// TIA Portal project "Vent Fan PLC" (V16) (continued)
VERSION : 0.1
   VAR_IN_OUT
      web_manual : "Station.Web_Interface.Manual.UDT";
      commands : "Drive.Commands.UDT";
   END_VAR
   VAR CONSTANT
      _RUN : String := 'run';
      _STOP : String := 'stop';
      _OVERRIDE : String := 'override';
   END_VAR
BEGIN
   "Drive.Commands.Run.Manual.Override"(web_manual := #web_manual,
                                        commands := #commands);
   IF #web_manual.mode <> #_OVERRIDE THEN
       "Drive.Commands.Run.Manual.Mode"(web_manual := #web_manual,
                                        commands := #commands);
   END_IF;
END_FUNCTION

FUNCTION "Schedule.In_Schedule" : Real   // FC11, SCL
{ S7_Optimized_Access := 'TRUE' }
VERSION : 0.1
   VAR_IN_OUT
      schedule : "Schedules.Temporal.UDT";
   END_VAR
   VAR_TEMP
      _now : DTL;
      _ret_val : Int;
      _monday : Real;
      _tuesday : Real;
      _wednesday : Real;
      _thursday : Real;
      _friday : Real;
      _saturday : Real;
      _sunday : Real;
   END_VAR
   // Ret_Val : returns speed if current time falls in any scheuled range
   VAR CONSTANT
      SUNDAY : USInt := 1;
      MONDAY : USInt := 2;
      TUESDAY : USInt := 3;
      WEDNESDAY : USInt := 4;
      THURSDAY : USInt := 5;
      FRIDAY : USInt := 6;
      SATURDAY : USInt := 7;
   END_VAR
BEGIN
   #_ret_val := RD_SYS_T(#_now);
   #_now.YEAR := 1970;
   #_now.HOUR -= 5;

   "Schedule.Encode_Weekday"(weekday := #MONDAY,
                             day_schedule := #schedule.monday);
   #_monday := "Schedule.In_Day"(day_schedule := #schedule.monday,
                                 current_time := #_now);
   IF #_monday > 0.0 THEN
       #"Schedule.In_Schedule" := #_monday;
       RETURN;
   END_IF;

   "Schedule.Encode_Weekday"(weekday := #TUESDAY,
                             day_schedule := #schedule.tuesday);
   #_tuesday := "Schedule.In_Day"(day_schedule := #schedule.tuesday,
                                  current_time := #_now);
   IF #_tuesday > 0.0 THEN
       #"Schedule.In_Schedule" := #_tuesday;
       RETURN;
   END_IF;

   "Schedule.Encode_Weekday"(weekday := #WEDNESDAY,
                             day_schedule := #schedule.wednesday);
   #_wednesday := "Schedule.In_Day"(day_schedule := #schedule.wednesday,
                                    current_time := #_now);
   IF #_wednesday > 0.0 THEN
       #"Schedule.In_Schedule" := #_wednesday;
       RETURN;
   END_IF;

   "Schedule.Encode_Weekday"(weekday := #THURSDAY,
                             day_schedule := #schedule.thursday);
   #_thursday := "Schedule.In_Day"(day_schedule := #schedule.thursday,
                                   current_time := #_now);
   IF #_thursday > 0.0 THEN
       #"Schedule.In_Schedule" := #_thursday;
       RETURN;
   END_IF;

   "Schedule.Encode_Weekday"(weekday := #FRIDAY,
                             day_schedule := #schedule.friday);
   #_friday := "Schedule.In_Day"(day_schedule := #schedule.friday,
                                 current_time := #_now);
   IF #_friday > 0.0 THEN
       #"Schedule.In_Schedule" := #_friday;
       RETURN;
   END_IF;

   "Schedule.Encode_Weekday"(weekday := #SATURDAY,
                             day_schedule := #schedule.saturday);
   #_saturday := "Schedule.In_Day"(day_schedule := #schedule.saturday,
                                   current_time := #_now);
   IF #_saturday > 0.0 THEN
       #"Schedule.In_Schedule" := #_saturday;
       RETURN;
   END_IF;

   "Schedule.Encode_Weekday"(weekday := #SUNDAY,
                             day_schedule := #schedule.sunday);
   #_sunday := "Schedule.In_Day"(day_schedule := #schedule.sunday,
                                 current_time := #_now);
   IF #_sunday > 0.0 THEN
       #"Schedule.In_Schedule" := #_sunday;
       RETURN;
   END_IF;

   #"Schedule.In_Schedule" := 0.0;
END_FUNCTION

FUNCTION "Drive.Commands.Run" : Void   // FC12, SCL
{ S7_Optimized_Access := 'TRUE' }
VERSION : 0.1
   VAR_INPUT
      current_station : Int;
      selected_station : Int;
      sensor : "Sensors.Thermal.UDT";
   END_VAR
   VAR_IN_OUT
      commands : "Drive.Commands.UDT";
      commands_manual : "Drive.Commands.UDT";
      commands_temporal : "Drive.Commands.UDT";
      commands_thermal : "Drive.Commands.UDT";
      web_manual : "Station.Web_Interface.Manual.UDT";
      thermal : "Schedules.Thermal.UDT";
      temporal : "Schedules.Temporal.UDT";
   END_VAR
BEGIN
   REGION "TEMPORAL"
       "Drive.Commands.Run.Temporal"(schedule:=#temporal,
                                     commands:=#commands_temporal);
       "Drive.Commands.Run.Temporal"(commands:=#commands_temporal,
                                     schedule:=#temporal);

   END_REGION

   REGION "THERMAL"
       "Drive.Commands.Run.Thermal"(sensor := #sensor,
                                    schedule := #thermal,
                                    commands := #commands_thermal);
   END_REGION

   REGION "MANUAL"
       IF #selected_station = #current_station THEN
           "Drive.Commands.Run.Manual"(web_manual := #web_manual,
                                       commands := #commands_manual);
       END_IF;
   END_REGION

   REGION "RESOLVE COMMANDS"
       "Drive.Commands.Run.Actual"(manual := #commands_manual,
                                   temporal := #commands_temporal,
                                   thermal := #commands_thermal,
                                   actual := #commands);
   END_REGION ;
END_FUNCTION

FUNCTION "Drive.Commands" : Void   // FC13, SCL
{ S7_Optimized_Access := 'TRUE' }
VERSION : 0.1
   VAR_INPUT
      current_station : Int;
      selected_station : Int;
      thermal_sensor : "Sensors.Thermal.UDT";
   END_VAR
   VAR_IN_OUT
      commands : "Drive.Commands.UDT";
      commands_manual : "Drive.Commands.UDT";
      commands_temporal : "Drive.Commands.UDT";
      commands_thermal : "Drive.Commands.UDT";
      manual : "Station.Web_Interface.Manual.UDT";
      thermal : "Schedules.Thermal.UDT";
      temporal : "Schedules.Temporal.UDT";
   END_VAR
BEGIN
   "Drive.Commands.Run"(current_station := #current_station,
                        selected_station := #selected_station,
                        sensor := #thermal_sensor,
                        commands := #commands,
                        commands_manual := #commands_manual,
                        commands_thermal := #commands_thermal,
                        commands_temporal := #commands_temporal,
                        web_manual := #manual,
                        thermal := #thermal,
                        temporal := #temporal);
END_FUNCTION

FUNCTION "Drive.Commands.Run.Actual" : Void   // FC14, SCL
{ S7_Optimized_Access := 'TRUE' }
VERSION : 0.1
   VAR_INPUT
      manual : "Drive.Commands.UDT";
      temporal : "Drive.Commands.UDT";
      thermal : "Drive.Commands.UDT";
   END_VAR
   VAR_IN_OUT
      actual : "Drive.Commands.UDT";
   END_VAR
BEGIN
   IF #manual.stop THEN
       #actual := #manual;
       RETURN;
   END_IF;

   IF #manual.override THEN
       #actual := #manual;
       RETURN;
   END_IF;

   IF #thermal.run THEN
       #actual := #thermal;
       RETURN;
   END_IF;

   IF #temporal.run THEN
       #actual := #temporal;
       RETURN;
   END_IF;

   #actual.speed := "Drive.Protection.Bound_Percentage"(#actual.speed);

   "Drive.Command_Stop"(#actual);
END_FUNCTION

FUNCTION "Real.Scale" : Real   // FC15, SCL
{ S7_Optimized_Access := 'TRUE' }
VERSION : 0.1
   VAR_INPUT
      x_min : Real;
      x_max : Real;
      x_actual : Real;
      y_min : Real;
      y_max : Real;
   END_VAR
BEGIN
   #"Real.Scale" := (#y_max - #y_min) / (#x_max - #x_min) * (#x_actual - #x_min) + (#y_min);
END_FUNCTION

FUNCTION "String.Split" : Void   // FC16, SCL
{ S7_Optimized_Access := 'TRUE' }
VERSION : 0.1
   VAR_INPUT
      string_in : String;
      delimeter : String;
      pointer : Int;   // pointer for recursion
   END_VAR
   VAR_IN_OUT
      sub_strings : Array[*] of String;
   END_VAR
   VAR_TEMP
      _split : String;
      _position : Int;
      _return : String;
   END_VAR
BEGIN
   REGION "GET POSITION OF DELIMETER IN STRING"
       #_position := FIND(IN1 := #string_in,
                          IN2 := #delimeter);
   END_REGION

   REGION "BASE CASE"
       IF #_position = 0 THEN
           #sub_strings[#pointer] := #string_in;
           RETURN;
       END_IF;
   END_REGION


   REGION "RECURSIVE CASE"
       #sub_strings[#pointer] := LEFT(IN := #string_in, L := #_position - 1);
       "String.Split"(string_in := RIGHT(IN := #string_in, L := LEN(#string_in) - #_position),
                      delimeter := #delimeter,
                      "pointer" := #pointer + 1,
                      sub_strings := #sub_strings);
   END_REGION
END_FUNCTION

FUNCTION "Schedule.Temporal.Clean_Data" : Void   // FC17, SCL
{ S7_Optimized_Access := 'TRUE' }
VERSION : 0.1
   VAR_IN_OUT
      schedule : "Schedules.Temporal.UDT";
   END_VAR
BEGIN
END_FUNCTION

FUNCTION "Web_Meta.Update_Temporal" : Void   // FC18, SCL
{ S7_Optimized_Access := 'TRUE' }
VERSION : 0.1
   VAR_IN_OUT
      web_schedules : "Web_Meta.Web_Interface.Schedules.Temporal.UDT";
      plc_schedules : "Schedules.Temporal.UDT";
   END_VAR
BEGIN
   IF NOT #web_schedules.new_data THEN
       RETURN;
   END_IF;

   "Web_Meta.Update_Temporal.Web_to_PLC"(web := #web_schedules,
                                         plc := #plc_schedules);
   #web_schedules.new_data := FALSE;
END_FUNCTION

FUNCTION "Web_Meta.Update_Temporal.Web_to_PLC" : Void   // FC19, SCL
{ S7_Optimized_Access := 'TRUE' }
VERSION : 0.1
   VAR_INPUT
      web : "Web_Meta.Web_Interface.Schedules.Temporal.UDT";
   END_VAR
   VAR_IN_OUT
      plc : "Schedules.Temporal.UDT";
   END_VAR
BEGIN
   "Web_Meta.Update_Temporal.Web_to_PLC.Day"(web := #web.monday,
                                             plc := #plc.monday);
   "Web_Meta.Update_Temporal.Web_to_PLC.Day"(web := #web.tuesday,
                                             plc := #plc.tuesday);
   "Web_Meta.Update_Temporal.Web_to_PLC.Day"(web := #web.wednesday,
                                             plc := #plc.wednesday);
   "Web_Meta.Update_Temporal.Web_to_PLC.Day"(web := #web.thursday,
                                             plc := #plc.thursday);
   "Web_Meta.Update_Temporal.Web_to_PLC.Day"(web := #web.friday,
                                             plc := #plc.friday);
   "Web_Meta.Update_Temporal.Web_to_PLC.Day"(web := #web.saturday,
                                             plc := #plc.saturday);
   "Web_Meta.Update_Temporal.Web_to_PLC.Day"(web := #web.sunday,
                                             plc := #plc.sunday);
END_FUNCTION

FUNCTION "Web_Meta.Update_Temporal.PLC_to_Web" : Void   // FC20, SCL
{ S7_Optimized_Access := 'TRUE' }
VERSION : 0.1
   VAR_INPUT
      plc : "Schedules.Temporal.UDT";
   END_VAR
   VAR_IN_OUT
      web : "Web_Meta.Web_Interface.Schedules.Temporal.UDT";
   END_VAR
BEGIN
   "Web_Meta.Update_Temporal.PLC_to_Web.Day"(plc := #plc.monday,
                                             web := #web.monday);
   "Web_Meta.Update_Temporal.PLC_to_Web.Day"(plc := #plc.tuesday,
                                             web := #web.tuesday);
   "Web_Meta.Update_Temporal.PLC_to_Web.Day"(plc := #plc.wednesday,
                                             web := #web.wednesday);
   "Web_Meta.Update_Temporal.PLC_to_Web.Day"(plc := #plc.thursday,
                                             web := #web.thursday);
   "Web_Meta.Update_Temporal.PLC_to_Web.Day"(plc := #plc.friday,
                                             web := #web.friday);
   "Web_Meta.Update_Temporal.PLC_to_Web.Day"(plc := #plc.saturday,
                                             web := #web.saturday);
   "Web_Meta.Update_Temporal.PLC_to_Web.Day"(plc := #plc.sunday,
                                             web := #web.sunday);
END_FUNCTION

FUNCTION "Web_Meta.Update_Temporal.PLC_to_Web.Day" : Void   // FC21, SCL
{ S7_Optimized_Access := 'TRUE' }
VERSION : 0.1
   VAR_INPUT
      plc : Array[0.."SCHEDULES_PER_DAY"] of "Schedules.Temporal.Element.UDT";
   END_VAR
   VAR_IN_OUT
      web : Array[0.."SCHEDULES_PER_DAY"] of "Web_Meta.Web_Interface.Schedules.Temporal.Element.UDT";
   END_VAR
   VAR_TEMP
      _i : Int;
   END_VAR
BEGIN
   FOR #_i := 0 TO "SCHEDULES_PER_DAY" DO
       #web[#_i].start := "Web_Meta.Update_Temporal.PLC_to_Web.Day.Element"(#plc[#_i].start);
       #web[#_i].stop := "Web_Meta.Update_Temporal.PLC_to_Web.Day.Element"(#plc[#_i].stop);
       #web[#_i].speed := #plc[#_i].speed;
   END_FOR;
END_FUNCTION

FUNCTION "Web_Meta.Update_Temporal.PLC_to_Web.Day.Element" : String   // FC22, SCL
{ S7_Optimized_Access := 'TRUE' }
VERSION : 0.1
   VAR_INPUT
      plc : "Schedules.Temporal.Element.Date_Time.UDT";
   END_VAR
   VAR_TEMP
      _ret : String;
   END_VAR
   VAR CONSTANT
      YEAR : String := '2022';
      "-" : String := '-';
   END_VAR
BEGIN
   // format --> value="2017-06-01T08:30"
   #_ret := CONCAT_STRING(IN1 := #YEAR,
                          IN2 := '-',
                          IN3 := "USInt.Convert.String.Date_with_Leading_Zeros"(#plc.month),
                          IN4 := '-',
                          IN5 := "USInt.Convert.String.Date_with_Leading_Zeros"(#plc.day),
                          IN6 := 'T',
                          IN7 := "USInt.Convert.String.Date_with_Leading_Zeros"(#plc.hour),
                          IN8 := ':',
                          IN9 := "USInt.Convert.String.Date_with_Leading_Zeros"(#plc.minute));
   #"Web_Meta.Update_Temporal.PLC_to_Web.Day.Element" := #_ret;
END_FUNCTION

FUNCTION "String.Strip Sign" : String   // FC23, SCL
{ S7_Optimized_Access := 'TRUE' }
VERSION : 0.1
   VAR_INPUT
      "string" : String;
   END_VAR
   VAR_TEMP
      Length : Int;
      "String Box" : String;
      "Test Character" : String;
   END_VAR
   VAR CONSTANT
      "+" : Char := '+';
      "-" : Char := '-';
   END_VAR
BEGIN
   #"String Box" := #string;
   #"Test Character" := LEFT_STRING(IN := #"String Box",
                                    L := 1);
   IF #"Test Character" = #"+" OR #"Test Character" = #"-" THEN
       #Length := LEN(#"String Box");
       #"String Box" := RIGHT_STRING(IN := #"String Box", L := #Length - 1);

   END_IF;
   #"String.Strip Sign" := #"String Box";
END_FUNCTION

FUNCTION "String.Trim" : String   // FC24, SCL
{ S7_Optimized_Access := 'TRUE' }
AUTHOR : Machado
FAMILY : String
VERSION : 1.0
// removes leading and trailing whitespace from input string
   VAR_INPUT
      "string" : String;
   END_VAR
   VAR_TEMP
      ret : String;
   END_VAR
   VAR CONSTANT
      space : String := ' ';
   END_VAR
BEGIN
   #ret := #string;
   WHILE LEFT(IN := #ret, L := 1) = #space DO
       #ret := RIGHT(IN := #ret, L := LEN(#ret) - 1);
   END_WHILE;
   WHILE RIGHT(IN := #ret, L := 1) = #space DO
       #ret := LEFT(IN := #ret, L := LEN(#ret) - 1);
   END_WHILE;
   #"String.Trim" := #ret;
END_FUNCTION

FUNCTION "USInt.Convert.Clean_String" : String   // FC25, SCL
{ S7_Optimized_Access := 'TRUE' }
VERSION : 0.1
   VAR_INPUT
      in : USInt;
   END_VAR
BEGIN
   #"USInt.Convert.Clean_String" := "String.Trim"("String.Strip Sign"(USINT_TO_STRING(#in)));
END_FUNCTION

FUNCTION "String.Add Leading" : String   // FC26, SCL
{ S7_Optimized_Access := 'TRUE' }
VERSION : 0.1
   VAR_INPUT
      "Leading Character" : Char;
      "Desired Length" : USInt;
      "String" : String;
   END_VAR
   VAR_TEMP
      Length : Int;
      "String Box" : String;
   END_VAR
BEGIN
   #"String Box" := #String;
   #Length := LEN(#"String Box");

   WHILE #Length < #"Desired Length" DO
       #"String Box" := CONCAT_STRING(IN1 := #"Leading Character",
                                      IN2 := #"String Box");
       #Length := LEN(#"String Box");
   END_WHILE;

   #"String.Add Leading" := #"String Box";
END_FUNCTION

FUNCTION "USInt.Convert.String.Date_with_Leading_Zeros" : String   // FC27, SCL
{ S7_Optimized_Access := 'TRUE' }
VERSION : 0.1
   VAR_INPUT
      in : USInt;
   END_VAR
BEGIN
   #"USInt.Convert.String.Date_with_Leading_Zeros" := "String.Add Leading"("Leading Character" := '0',
                                                                           "Desired Length" := 2,
                                                                           "String" := "USInt.Convert.Clean_String"(#in));
END_FUNCTION

FUNCTION "Web_Meta.Update_Temporal.Web_to_PLC.Day.Element" : "Schedules.Temporal.Element.Date_Time.UDT"   // FC28, SCL
{ S7_Optimized_Access := 'TRUE' }
VERSION : 0.1
   VAR_INPUT
      in : String;
   END_VAR
   VAR_TEMP
      _ret : "Schedules.Temporal.Element.Date_Time.UDT";
      _split_date_time : Array[0..1] of String;
      _split_date : Array[0..2] of String;
      _split_time : Array[0..1] of String;
   END_VAR
BEGIN
   // format --> value="2017-06-01T08:30"
   REGION "SPLIT INTO DATE AND TIME"
       "String.Split"(string_in := #in,
                      delimeter := 'T',
                      "pointer" := 0,
                      sub_strings := #_split_date_time);
   END_REGION

   REGION "SPLIT DATE INTO YEARS, MONTHS, AND DAYS"
       "String.Split"(string_in := #_split_date_time[0],
                      delimeter := '-',
                      "pointer" := 0,
                      sub_strings := #_split_date);
   END_REGION

   REGION "SPLIT TIME INTO HOURS AND MINUTES"
       "String.Split"(string_in := #_split_date_time[1],
                      delimeter := ':',
                      "pointer" := 0,
                      sub_strings := #_split_time);
   END_REGION

   REGION "MAP TO UDT"
       #_ret.month := STRING_TO_USINT(#_split_date[1]);
       #_ret.day := STRING_TO_USINT(#_split_date[2]);
       #_ret.hour := STRING_TO_USINT(#_split_time[0]);
       #_ret.minute := STRING_TO_USINT(#_split_time[1]);
   END_REGION

   REGION "RETURN DATA"
       #"Web_Meta.Update_Temporal.Web_to_PLC.Day.Element" := #_ret;
   END_REGION
END_FUNCTION

FUNCTION "Web_Meta.Update_Temporal.Web_to_PLC.Day" : Void   // FC29, SCL
{ S7_Optimized_Access := 'TRUE' }
VERSION : 0.1
   VAR_INPUT
      web : Array[0.."SCHEDULES_PER_DAY"] of "Web_Meta.Web_Interface.Schedules.Temporal.Element.UDT";
   END_VAR
   VAR_IN_OUT
      plc : Array[0.."SCHEDULES_PER_DAY"] of "Schedules.Temporal.Element.UDT";
   END_VAR
   VAR_TEMP
      _i : Int;
   END_VAR
BEGIN
   FOR #_i := 0 TO "SCHEDULES_PER_DAY" DO
       #plc[#_i].start := "Web_Meta.Update_Temporal.Web_to_PLC.Day.Element"(#web[#_i].start);
       #plc[#_i].stop := "Web_Meta.Update_Temporal.Web_to_PLC.Day.Element"(#web[#_i].stop);
       #plc[#_i].speed := #web[#_i].speed;
   END_FOR;
END_FUNCTION

FUNCTION "Schedule.In_Day" : Real   // FC30, SCL
{ S7_Optimized_Access := 'TRUE' }
VERSION : 0.1
   VAR_INPUT
      day_schedule : Array[0.."SCHEDULES_PER_DAY"] of "Schedules.Temporal.Element.UDT";
      current_time : DTL;
   END_VAR
   VAR_TEMP
      _i : Int;
      _speed : Real;
   END_VAR
BEGIN
   IF #current_time.WEEKDAY <> #day_schedule[0].start.weekday THEN
       #"Schedule.In_Day" := 0.0;
       RETURN;
   END_IF;
   FOR #_i := 0 TO "SCHEDULES_PER_DAY" DO
       #_speed := "Schedule.In_Window"(day := #day_schedule[#_i],
                                       now := #current_time);
       IF #_speed > 0.0 THEN
           #"Schedule.In_Day" := #_speed;
           RETURN;
       END_IF;
   END_FOR;
   #"Schedule.In_Day" := 0.0;
END_FUNCTION

FUNCTION "Schedule.In_Window" : Real   // FC31, SCL
{ S7_Optimized_Access := 'TRUE' }
VERSION : 0.1
   VAR_INPUT
      day : "Schedules.Temporal.Element.UDT";
      now : DTL;
   END_VAR
   VAR_TEMP
      _start : DTL;
      _stop : DTL;
   END_VAR
BEGIN
   #_start := "Schedule.Map.Date_Time_to_DTL"(#day.start);
   #_stop := "Schedule.Map.Date_Time_to_DTL"(#day.stop);
   IF #_start < #now AND #now < #_stop THEN
       #"Schedule.In_Window" := #day.speed;
       RETURN;
   END_IF;
   #"Schedule.In_Window" := 0.0;
END_FUNCTION

FUNCTION "Schedule.Map.Date_Time_to_DTL" : DTL   // FC32, SCL
{ S7_Optimized_Access := 'TRUE' }
VERSION : 0.1
   VAR_INPUT
      boundary : "Schedules.Temporal.Element.Date_Time.UDT";
   END_VAR
   VAR_TEMP
      _ret : DTL;
   END_VAR
BEGIN
   #_ret.MONTH := #boundary.month;
   #_ret.DAY := #boundary.day;
   #_ret.HOUR := #boundary.hour;
   #_ret.MINUTE := #boundary.minute;
   #"Schedule.Map.Date_Time_to_DTL" := #_ret;
END_FUNCTION

FUNCTION "Drive.Commands.Run.Temporal" : Void   // FC33, SCL
{ S7_Optimized_Access := 'TRUE' }
VERSION : 0.1
   VAR_IN_OUT
      commands : "Drive.Commands.UDT";
      schedule : "Schedules.Temporal.UDT";
   END_VAR
   VAR_TEMP
      _speed : Real;
   END_VAR
BEGIN
   #_speed := "Schedule.In_Schedule"(schedule:=#schedule);

   IF #_speed = 0.0 THEN
       "Drive.Command_Stop"(#commands);
       RETURN;
   END_IF;

   "Drive.Command_Run"(speed := #_speed,
                       commands := #commands);
END_FUNCTION

FUNCTION "Drive.Command_Run" : Void   // FC34, SCL
{ S7_Optimized_Access := 'TRUE' }
VERSION : 0.1
   VAR_INPUT
      speed : Real;
   END_VAR
   VAR_IN_OUT
      commands : "Drive.Commands.UDT";
   END_VAR
BEGIN
   #commands.run := TRUE;
   #commands.stop := FALSE;
   #commands.speed := #speed;
END_FUNCTION

FUNCTION "Drive.Command_Stop" : Void   // FC35, SCL
{ S7_Optimized_Access := 'TRUE' }
VERSION : 0.1
   VAR_IN_OUT
      commands : "Drive.Commands.UDT";
   END_VAR
BEGIN
   #commands.run := FALSE;
   #commands.stop := TRUE;
   #commands.speed := 0.0;
END_FUNCTION

FUNCTION "Nibble.ToString" : String   // FC36, SCL
{ S7_Optimized_Access := 'TRUE' }
VERSION : 0.1
   VAR_INPUT
      value : Byte;
   END_VAR
   VAR_TEMP
      _nibble_as_int : Int;
      _ret : String;
   END_VAR
BEGIN
   #_nibble_as_int := BYTE_TO_INT(#value);
   CASE #_nibble_as_int OF
       0..9:
           #_ret := "String.Trim"("String.Strip Sign"(INT_TO_STRING(#_nibble_as_int)));
       10:
           #_ret := 'A';
       11:
           #_ret := 'B';
       12:
           #_ret := 'C';
       13:
           #_ret := 'D';
       14:
           #_ret := 'E';
       15:
           #_ret := 'F';
   END_CASE;
   #"Nibble.ToString" := #_ret;
END_FUNCTION

FUNCTION "Byte.ToString" : String   // FC37, SCL
{ S7_Optimized_Access := 'TRUE' }
VERSION : 0.1
   VAR_INPUT
      value : Byte;
   END_VAR
   VAR_TEMP
      _low_nibble : Byte;
      _high_nibble : Byte;
   END_VAR
   VAR CONSTANT
      LOW_NIBBLE_MASK : Byte := 16#0F;
      HIGH_NIBBLE_MASK : Byte := 16#F0;
   END_VAR
BEGIN
   #_low_nibble := #value AND #LOW_NIBBLE_MASK;
   #_high_nibble := SHR_BYTE(IN := #value AND #HIGH_NIBBLE_MASK,
                             N := 4);
   #"Byte.ToString" := CONCAT_STRING(IN1 := "Nibble.ToString"(#_high_nibble),
                                     IN2 := "Nibble.ToString"(#_low_nibble));
END_FUNCTION

FUNCTION "Drive.Feedback.Speed.Percent_to_RPM" : Real   // FC38, SCL
{ S7_Optimized_Access := 'TRUE' }
VERSION : 0.1
   VAR_INPUT
      as_percent : Real;
      max_speed : Real;
   END_VAR
BEGIN
   #"Drive.Feedback.Speed.Percent_to_RPM" := "Drive.Protection.Bound_Percentage"(#as_percent/100) * #max_speed;
END_FUNCTION

FUNCTION "Drive.Protection.Bound_Percentage" : Real   // FC39, SCL
{ S7_Optimized_Access := 'TRUE' }
VERSION : 0.1
   VAR_INPUT
      value : Real;
   END_VAR
BEGIN
   IF #value > 1.0 THEN
       #"Drive.Protection.Bound_Percentage" := 1.0;
       RETURN;
   END_IF;

   IF #value < 0.0 THEN
       #"Drive.Protection.Bound_Percentage" := 0.0;
       RETURN;
   END_IF;

   #"Drive.Protection.Bound_Percentage" := #value;
END_FUNCTION

FUNCTION "Schedule.Encode_Weekday" : Void   // FC40, SCL
{ S7_Optimized_Access := 'TRUE' }
VERSION : 0.1
   VAR_INPUT
      weekday : USInt;
   END_VAR
   VAR_IN_OUT
      day_schedule : Array[0.."SCHEDULES_PER_DAY"] of "Schedules.Temporal.Element.UDT";
   END_VAR
   VAR_TEMP
      i : Int;
   END_VAR
BEGIN
   FOR #i := 0 TO "SCHEDULES_PER_DAY" DO
       #day_schedule[#i].start.weekday := #weekday;
       #day_schedule[#i].stop.weekday := #weekday;
   END_FOR;
END_FUNCTION

FUNCTION "Drive.Feedback.Speed.RPM_to_Percent" : Real   // FC41, SCL
{ S7_Optimized_Access := 'TRUE' }
VERSION : 0.1
   VAR_INPUT
      as_rpm : Real;
      max_speed : Real;
   END_VAR
BEGIN
   #"Drive.Feedback.Speed.RPM_to_Percent" := #as_rpm / #max_speed * 100.0;
END_FUNCTION

FUNCTION "Drive.Commands.Run.Manual.Override" : Void   // FC42, SCL
{ S7_Optimized_Access := 'TRUE' }
VERSION : 0.1
   VAR_IN_OUT
      web_manual : "Station.Web_Interface.Manual.UDT";
      commands : "Drive.Commands.UDT";
   END_VAR
   VAR CONSTANT
      _RUN : String := 'run';
      _STOP : String := 'stop';
      _OVERRIDE : String := 'override';
   END_VAR
BEGIN
   IF #web_manual.toggle AND #web_manual.mode = #_OVERRIDE THEN
       #web_manual.mode := #_STOP;
       #web_manual.toggle := FALSE;
       #web_manual.override := FALSE;
       #commands.override := FALSE;
       #commands.run := FALSE;
       #commands.stop := TRUE;
       #commands.speed := 0.0;
       RETURN;
   END_IF;
   IF #web_manual.override THEN
       #web_manual.mode := #_OVERRIDE;
       #commands.override := TRUE;
       #commands.run := TRUE;
       #commands.stop := FALSE;
       #commands.speed := #web_manual.command_speed;
       RETURN;
   END_IF;
   IF NOT #web_manual.override AND #web_manual.mode = #_OVERRIDE THEN
       #web_manual.mode := #_STOP;
       #commands.override := FALSE;
       #commands.run := FALSE;
       #commands.stop := TRUE;
       #commands.speed := 0.0;
   END_IF;
END_FUNCTION

FUNCTION "Drive.Commands.Run.Manual.Mode" : Void   // FC43, SCL
{ S7_Optimized_Access := 'TRUE' }
VERSION : 0.1
   VAR_IN_OUT
      web_manual : "Station.Web_Interface.Manual.UDT";
      commands : "Drive.Commands.UDT";
   END_VAR
   VAR CONSTANT
      _RUN : String := 'run';
      _STOP : String := 'stop';
   END_VAR
BEGIN
   IF NOT #web_manual.toggle THEN
       RETURN;
   END_IF;
   IF #web_manual.mode = #_RUN THEN
       #web_manual.mode := #_STOP;
       #commands.run := FALSE;
       #commands.stop := TRUE;
       #commands.speed := 0.0;
       #web_manual.toggle := FALSE;
       RETURN;
   END_IF;
   IF #web_manual.mode = #_STOP THEN
       #web_manual.mode := #_RUN;
       #commands.run := TRUE;
       #commands.stop := FALSE;
       #web_manual.toggle := FALSE;
   END_IF;
END_FUNCTION

FUNCTION "Web_Meta.Update_Manual.PLC_to_Web" : Void   // FC44, SCL
{ S7_Optimized_Access := 'TRUE' }
VERSION : 0.1
   VAR_INPUT
      station : "Station.UDT";
   END_VAR
   VAR_IN_OUT
      manual : "Station.Web_Interface.Manual.UDT";
   END_VAR
BEGIN
   #manual.command_speed := #station.drive.commands_manual.speed;
   #manual.override := #station.drive.commands_manual.override;
   IF #station.drive.commands.override THEN
       #manual.mode := 'override';
   END_IF;
   IF #station.drive.commands.run THEN
       #manual.mode := 'run';
   END_IF;
   IF #station.drive.commands.stop THEN
       #manual.mode := 'stop';
   END_IF;
END_FUNCTION

FUNCTION "Faults" : Void   // FC45, SCL
{ S7_Optimized_Access := 'TRUE' }
VERSION : 0.1
   VAR_INPUT
      fault_code : Word;
   END_VAR
   VAR_IN_OUT
      station : "Station.UDT";
   END_VAR
   VAR_TEMP
      _drive_speed : Real;
      _command_speed : Real;
      _current : Real;
   END_VAR
   VAR CONSTANT
      NO_FAULT : Word := 16#7002;
      COMM_FAULT : Word := 16#80B1;
      RED : String := 'red';
      BLUE : String := 'blue';
      YELLOW : String := 'yellow';
      GREEN : String := 'green';
   END_VAR
BEGIN
   #station.faults.fault := 'no faults';
   #station.faults.color := '';

   #_drive_speed := #station.drive.feedback.speed.me.processed;
   #_command_speed := #station.drive.commands.speed;
   #_current := #station.drive.feedback.current.me.processed;

   IF #fault_code >= #NO_FAULT THEN
       IF #fault_code <> #COMM_FAULT THEN
           #station.faults.fault := "Word.ToString"(#fault_code);
           #station.faults.color := #RED;
           RETURN;
       END_IF;
   END_IF;

   IF #_drive_speed = 0.0 THEN
       IF #_command_speed <> 0.0 THEN
           #station.faults.fault := 'stopped while commanded speed above 0.0';
           #station.faults.color := #YELLOW;
           RETURN;
       END_IF;
   END_IF;

   IF #_command_speed > 10.0 THEN
       IF #_current < 2.0 THEN
           #station.faults.fault := 'low current draw';
           #station.faults.color := #RED;
           RETURN;
       END_IF;
   END_IF;

   IF #_command_speed > 10.0 THEN
       IF #_current > 6.0 THEN
           #station.faults.fault := 'high current draw';
           #station.faults.color := #RED;
           RETURN;
       END_IF;
   END_IF;

   IF #_current > 7.0 THEN
       #station.drive.commands.speed := 0.0;
       #station.faults.fault := 'over current';
       #station.faults.color := #RED;
       RETURN;
   END_IF;

   IF #_drive_speed = 0.0 THEN
       IF #_command_speed = 0.0 THEN
           #station.faults.fault := 'drive commanded stop';
           #station.faults.color := #BLUE;
           RETURN;
       END_IF;
   END_IF;

   IF #_drive_speed > 0.9 * #_command_speed THEN
       IF #_drive_speed < 1.1 * #_command_speed THEN
           #station.faults.fault := 'no faults';
           #station.faults.color := #GREEN;
           RETURN;
       END_IF;
   END_IF;
END_FUNCTION

ORGANIZATION_BLOCK "Main"   // OB1, LAD, ProgramCycle
TITLE = "Main Program Sweep (Cycle)"
{ S7_Optimized_Access := 'TRUE' }
VERSION : 0.1
   VAR_INPUT
      Initial_Call : Bool;   // Initial call of this OB
      Remanence : Bool;   // =True, if remanent data are available
   END_VAR
   VAR_TEMP
      RET_VAL : Int;
   END_VAR
   VAR CONSTANT
      SENSOR_MAX : Word := 16#3F_FF;
      SENSOR_MIN : Word;
      THERMAL_MAX : Real := 150.0;
      THERMAL_MIN : Real;
   END_VAR
BEGIN

REGION Network 1
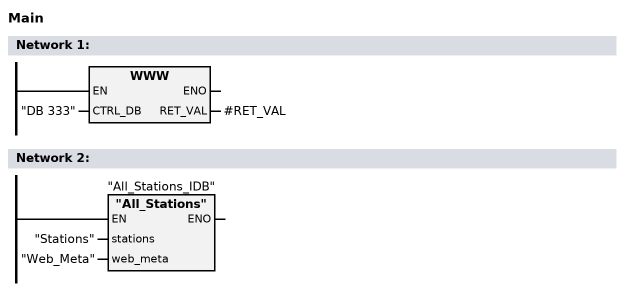
   #RET_VAL := WWW(CTRL_DB := "DB 333");
END_REGION

REGION Network 2
   RUNG wire#powerrail
      "All_Stations_IDB"(stations := "Stations", web_meta := "Web_Meta")
   END_RUNG
   // the same network as SCL:
   "All_Stations_IDB"(stations := "Stations", web_meta := "Web_Meta");   // "All_Stations"
END_REGION
END_ORGANIZATION_BLOCK

ORGANIZATION_BLOCK "Time error interrupt"   // OB80, LAD, TimeErrorInterrupt
{ S7_Optimized_Access := 'TRUE' }
VERSION : 0.1
   VAR_INPUT
      Fault_ID : Byte;   // Fault identifier
      Csg_OBnr : OB_Any;   // Number of OB causing the error
      Csg_Prio : UInt;   // Priority of OB causing the error
   END_VAR
BEGIN
END_ORGANIZATION_BLOCK